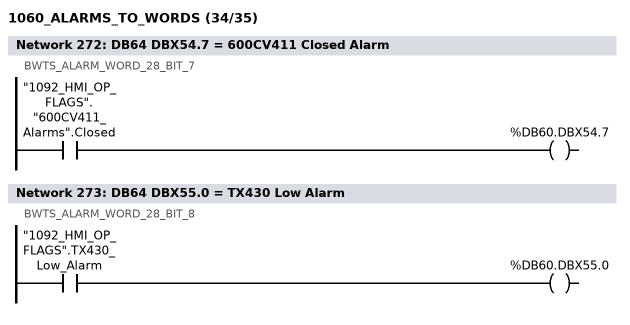
   RUNG wire#powerrail
      Contact( "1092_HMI_OP_FLAGS"."600CV411_Alarms".Closed )
      Coil( %DB60.DBX54.7 )
   END_RUNG
   // the same network as SCL:
   %DB60.DBX54.7 := "1092_HMI_OP_FLAGS"."600CV411_Alarms".Closed;
END_REGION

REGION Network 273: DB64 DBX55.0 = TX430 Low Alarm
   // BWTS_ALARM_WORD_28_BIT_8
   RUNG wire#powerrail
      Contact( "1092_HMI_OP_FLAGS".TX430_Low_Alarm )
      Coil( %DB60.DBX55.0 )
   END_RUNG
   // the same network as SCL:
   %DB60.DBX55.0 := "1092_HMI_OP_FLAGS".TX430_Low_Alarm;
END_REGION

REGION Network 275: Alarm Present
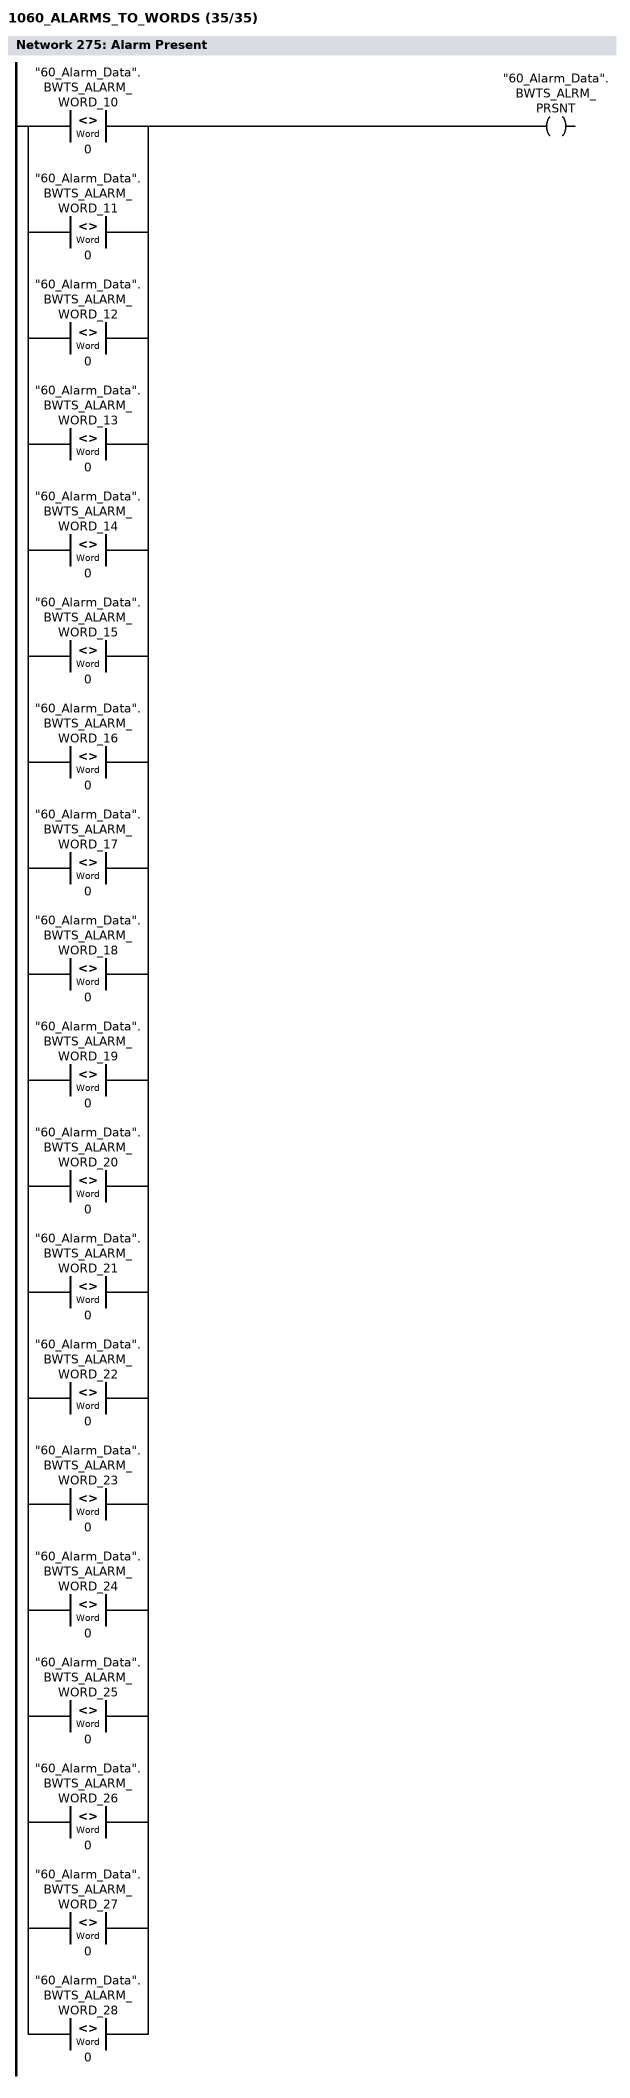
   RUNG wire#powerrail
      { S7_Templates := "SrcType := Word" } NE_Contact(in1 := "60_Alarm_Data".BWTS_ALARM_WORD_10, in2 := 0)
      wire#w1
      Coil( "60_Alarm_Data".BWTS_ALRM_PRSNT )
   END_RUNG
   RUNG wire#powerrail
      { S7_Templates := "SrcType := Word" } NE_Contact(in1 := "60_Alarm_Data".BWTS_ALARM_WORD_11, in2 := 0)
   END_RUNG wire#w1
   RUNG wire#powerrail
      { S7_Templates := "SrcType := Word" } NE_Contact(in1 := "60_Alarm_Data".BWTS_ALARM_WORD_12, in2 := 0)
   END_RUNG wire#w1
   RUNG wire#powerrail
      { S7_Templates := "SrcType := Word" } NE_Contact(in1 := "60_Alarm_Data".BWTS_ALARM_WORD_13, in2 := 0)
   END_RUNG wire#w1
   RUNG wire#powerrail
      { S7_Templates := "SrcType := Word" } NE_Contact(in1 := "60_Alarm_Data".BWTS_ALARM_WORD_14, in2 := 0)
   END_RUNG wire#w1
   RUNG wire#powerrail
      { S7_Templates := "SrcType := Word" } NE_Contact(in1 := "60_Alarm_Data".BWTS_ALARM_WORD_15, in2 := 0)
   END_RUNG wire#w1
   RUNG wire#powerrail
      { S7_Templates := "SrcType := Word" } NE_Contact(in1 := "60_Alarm_Data".BWTS_ALARM_WORD_16, in2 := 0)
   END_RUNG wire#w1
   RUNG wire#powerrail
      { S7_Templates := "SrcType := Word" } NE_Contact(in1 := "60_Alarm_Data".BWTS_ALARM_WORD_17, in2 := 0)
   END_RUNG wire#w1
   RUNG wire#powerrail
      { S7_Templates := "SrcType := Word" } NE_Contact(in1 := "60_Alarm_Data".BWTS_ALARM_WORD_18, in2 := 0)
   END_RUNG wire#w1
   RUNG wire#powerrail
      { S7_Templates := "SrcType := Word" } NE_Contact(in1 := "60_Alarm_Data".BWTS_ALARM_WORD_19, in2 := 0)
   END_RUNG wire#w1
   RUNG wire#powerrail
      { S7_Templates := "SrcType := Word" } NE_Contact(in1 := "60_Alarm_Data".BWTS_ALARM_WORD_20, in2 := 0)
   END_RUNG wire#w1
   RUNG wire#powerrail
      { S7_Templates := "SrcType := Word" } NE_Contact(in1 := "60_Alarm_Data".BWTS_ALARM_WORD_21, in2 := 0)
   END_RUNG wire#w1
   RUNG wire#powerrail
      { S7_Templates := "SrcType := Word" } NE_Contact(in1 := "60_Alarm_Data".BWTS_ALARM_WORD_22, in2 := 0)
   END_RUNG wire#w1
   RUNG wire#powerrail
      { S7_Templates := "SrcType := Word" } NE_Contact(in1 := "60_Alarm_Data".BWTS_ALARM_WORD_23, in2 := 0)
   END_RUNG wire#w1
   RUNG wire#powerrail
      { S7_Templates := "SrcType := Word" } NE_Contact(in1 := "60_Alarm_Data".BWTS_ALARM_WORD_24, in2 := 0)
   END_RUNG wire#w1
   RUNG wire#powerrail
      { S7_Templates := "SrcType := Word" } NE_Contact(in1 := "60_Alarm_Data".BWTS_ALARM_WORD_25, in2 := 0)
   END_RUNG wire#w1
   RUNG wire#powerrail
      { S7_Templates := "SrcType := Word" } NE_Contact(in1 := "60_Alarm_Data".BWTS_ALARM_WORD_26, in2 := 0)
   END_RUNG wire#w1
   RUNG wire#powerrail
      { S7_Templates := "SrcType := Word" } NE_Contact(in1 := "60_Alarm_Data".BWTS_ALARM_WORD_27, in2 := 0)
   END_RUNG wire#w1
   RUNG wire#powerrail
      { S7_Templates := "SrcType := Word" } NE_Contact(in1 := "60_Alarm_Data".BWTS_ALARM_WORD_28, in2 := 0)
   END_RUNG wire#w1
   // the same network as SCL:
   "60_Alarm_Data".BWTS_ALRM_PRSNT := ("60_Alarm_Data".BWTS_ALARM_WORD_10 <> 0) OR ("60_Alarm_Data".BWTS_ALARM_WORD_11 <> 0) OR ("60_Alarm_Data".BWTS_ALARM_WORD_12 <> 0) OR ("60_Alarm_Data".BWTS_ALARM_WORD_13 <> 0) OR ("60_Alarm_Data".BWTS_ALARM_WORD_14 <> 0) OR ("60_Alarm_Data".BWTS_ALARM_WORD_15 <> 0) OR ("60_Alarm_Data".BWTS_ALARM_WORD_16 <> 0) OR ("60_Alarm_Data".BWTS_ALARM_WORD_17 <> 0) OR ("60_Alarm_Data".BWTS_ALARM_WORD_18 <> 0) OR ("60_Alarm_Data".BWTS_ALARM_WORD_19 <> 0) OR ("60_Alarm_Data".BWTS_ALARM_WORD_20 <> 0) OR ("60_Alarm_Data".BWTS_ALARM_WORD_21 <> 0) OR ("60_Alarm_Data".BWTS_ALARM_WORD_22 <> 0) OR ("60_Alarm_Data".BWTS_ALARM_WORD_23 <> 0) OR ("60_Alarm_Data".BWTS_ALARM_WORD_24 <> 0) OR ("60_Alarm_Data".BWTS_ALARM_WORD_25 <> 0) OR ("60_Alarm_Data".BWTS_ALARM_WORD_26 <> 0) OR ("60_Alarm_Data".BWTS_ALARM_WORD_27 <> 0) OR ("60_Alarm_Data".BWTS_ALARM_WORD_28 <> 0);
END_REGION
END_FUNCTION

FUNCTION "1062_WARNINGS_TO_WORDS" : Void   // FC1062, LAD
TITLE = Warning Processing
{ S7_Optimized_Access := 'TRUE' }
AUTHOR : JRS
VERSION : 0.1
BEGIN

REGION Network 1: DB66 DBX18.0 = TX425/426 Tank 1 pH High Warning
   // BWTS_WARNING_WORD_10_BIT_0
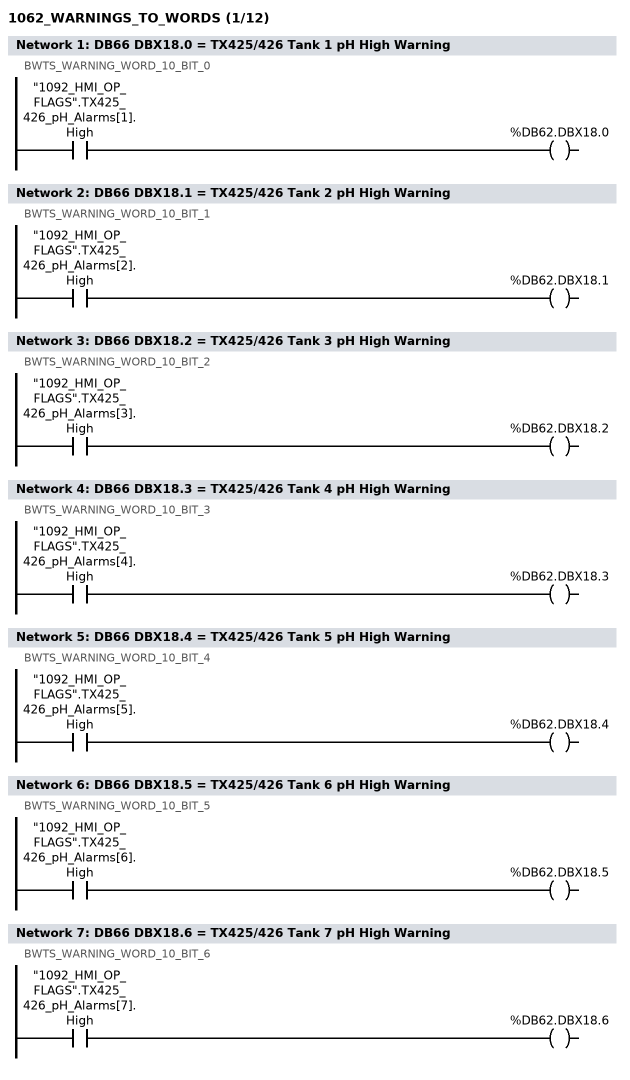
   RUNG wire#powerrail
      Contact( "1092_HMI_OP_FLAGS".TX425_426_pH_Alarms[1].High )
      Coil( %DB62.DBX18.0 )
   END_RUNG
   // the same network as SCL:
   %DB62.DBX18.0 := "1092_HMI_OP_FLAGS".TX425_426_pH_Alarms[1].High;
END_REGION

REGION Network 2: DB66 DBX18.1 = TX425/426 Tank 2 pH High Warning
   // BWTS_WARNING_WORD_10_BIT_1
   RUNG wire#powerrail
      Contact( "1092_HMI_OP_FLAGS".TX425_426_pH_Alarms[2].High )
      Coil( %DB62.DBX18.1 )
   END_RUNG
   // the same network as SCL:
   %DB62.DBX18.1 := "1092_HMI_OP_FLAGS".TX425_426_pH_Alarms[2].High;
END_REGION

REGION Network 3: DB66 DBX18.2 = TX425/426 Tank 3 pH High Warning
   // BWTS_WARNING_WORD_10_BIT_2
   RUNG wire#powerrail
      Contact( "1092_HMI_OP_FLAGS".TX425_426_pH_Alarms[3].High )
      Coil( %DB62.DBX18.2 )
   END_RUNG
   // the same network as SCL:
   %DB62.DBX18.2 := "1092_HMI_OP_FLAGS".TX425_426_pH_Alarms[3].High;
END_REGION

REGION Network 4: DB66 DBX18.3 = TX425/426 Tank 4 pH High Warning
   // BWTS_WARNING_WORD_10_BIT_3
   RUNG wire#powerrail
      Contact( "1092_HMI_OP_FLAGS".TX425_426_pH_Alarms[4].High )
      Coil( %DB62.DBX18.3 )
   END_RUNG
   // the same network as SCL:
   %DB62.DBX18.3 := "1092_HMI_OP_FLAGS".TX425_426_pH_Alarms[4].High;
END_REGION

REGION Network 5: DB66 DBX18.4 = TX425/426 Tank 5 pH High Warning
   // BWTS_WARNING_WORD_10_BIT_4
   RUNG wire#powerrail
      Contact( "1092_HMI_OP_FLAGS".TX425_426_pH_Alarms[5].High )
      Coil( %DB62.DBX18.4 )
   END_RUNG
   // the same network as SCL:
   %DB62.DBX18.4 := "1092_HMI_OP_FLAGS".TX425_426_pH_Alarms[5].High;
END_REGION

REGION Network 6: DB66 DBX18.5 = TX425/426 Tank 6 pH High Warning
   // BWTS_WARNING_WORD_10_BIT_5
   RUNG wire#powerrail
      Contact( "1092_HMI_OP_FLAGS".TX425_426_pH_Alarms[6].High )
      Coil( %DB62.DBX18.5 )
   END_RUNG
   // the same network as SCL:
   %DB62.DBX18.5 := "1092_HMI_OP_FLAGS".TX425_426_pH_Alarms[6].High;
END_REGION

REGION Network 7: DB66 DBX18.6 = TX425/426 Tank 7 pH High Warning
   // BWTS_WARNING_WORD_10_BIT_6
   RUNG wire#powerrail
      Contact( "1092_HMI_OP_FLAGS".TX425_426_pH_Alarms[7].High )
      Coil( %DB62.DBX18.6 )
   END_RUNG
   // the same network as SCL:
   %DB62.DBX18.6 := "1092_HMI_OP_FLAGS".TX425_426_pH_Alarms[7].High;
END_REGION

REGION Network 8: DB66 DBX18.7 = TX425/426 Tank 8 pH High Warning
   // BWTS_WARNING_WORD_10_BIT_7
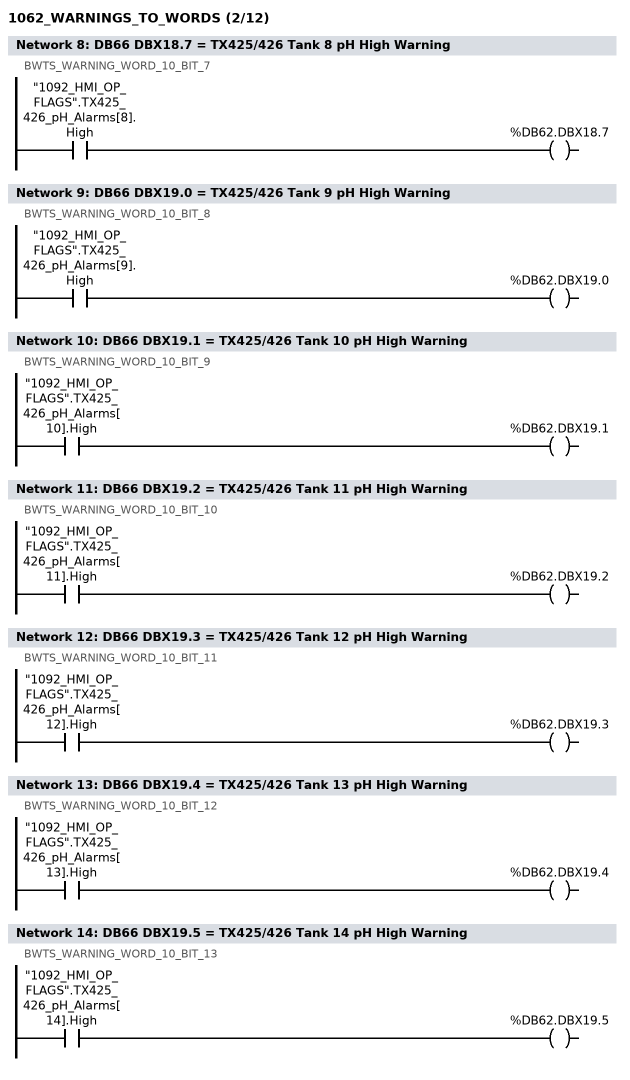
   RUNG wire#powerrail
      Contact( "1092_HMI_OP_FLAGS".TX425_426_pH_Alarms[8].High )
      Coil( %DB62.DBX18.7 )
   END_RUNG
   // the same network as SCL:
   %DB62.DBX18.7 := "1092_HMI_OP_FLAGS".TX425_426_pH_Alarms[8].High;
END_REGION

REGION Network 9: DB66 DBX19.0 = TX425/426 Tank 9 pH High Warning
   // BWTS_WARNING_WORD_10_BIT_8
   RUNG wire#powerrail
      Contact( "1092_HMI_OP_FLAGS".TX425_426_pH_Alarms[9].High )
      Coil( %DB62.DBX19.0 )
   END_RUNG
   // the same network as SCL:
   %DB62.DBX19.0 := "1092_HMI_OP_FLAGS".TX425_426_pH_Alarms[9].High;
END_REGION

REGION Network 10: DB66 DBX19.1 = TX425/426 Tank 10 pH High Warning
   // BWTS_WARNING_WORD_10_BIT_9
   RUNG wire#powerrail
      Contact( "1092_HMI_OP_FLAGS".TX425_426_pH_Alarms[10].High )
      Coil( %DB62.DBX19.1 )
   END_RUNG
   // the same network as SCL:
   %DB62.DBX19.1 := "1092_HMI_OP_FLAGS".TX425_426_pH_Alarms[10].High;
END_REGION

REGION Network 11: DB66 DBX19.2 = TX425/426 Tank 11 pH High Warning
   // BWTS_WARNING_WORD_10_BIT_10
   RUNG wire#powerrail
      Contact( "1092_HMI_OP_FLAGS".TX425_426_pH_Alarms[11].High )
      Coil( %DB62.DBX19.2 )
   END_RUNG
   // the same network as SCL:
   %DB62.DBX19.2 := "1092_HMI_OP_FLAGS".TX425_426_pH_Alarms[11].High;
END_REGION

REGION Network 12: DB66 DBX19.3 = TX425/426 Tank 12 pH High Warning
   // BWTS_WARNING_WORD_10_BIT_11
   RUNG wire#powerrail
      Contact( "1092_HMI_OP_FLAGS".TX425_426_pH_Alarms[12].High )
      Coil( %DB62.DBX19.3 )
   END_RUNG
   // the same network as SCL:
   %DB62.DBX19.3 := "1092_HMI_OP_FLAGS".TX425_426_pH_Alarms[12].High;
END_REGION

REGION Network 13: DB66 DBX19.4 = TX425/426 Tank 13 pH High Warning
   // BWTS_WARNING_WORD_10_BIT_12
   RUNG wire#powerrail
      Contact( "1092_HMI_OP_FLAGS".TX425_426_pH_Alarms[13].High )
      Coil( %DB62.DBX19.4 )
   END_RUNG
   // the same network as SCL:
   %DB62.DBX19.4 := "1092_HMI_OP_FLAGS".TX425_426_pH_Alarms[13].High;
END_REGION

REGION Network 14: DB66 DBX19.5 = TX425/426 Tank 14 pH High Warning
   // BWTS_WARNING_WORD_10_BIT_13
   RUNG wire#powerrail
      Contact( "1092_HMI_OP_FLAGS".TX425_426_pH_Alarms[14].High )
      Coil( %DB62.DBX19.5 )
   END_RUNG
   // the same network as SCL:
   %DB62.DBX19.5 := "1092_HMI_OP_FLAGS".TX425_426_pH_Alarms[14].High;
END_REGION

REGION Network 16: DB66 DBX20.0 = FIT417/418 Flow Tank 1 High Warning
   // BWTS_WARNING_WORD_11_BIT_0
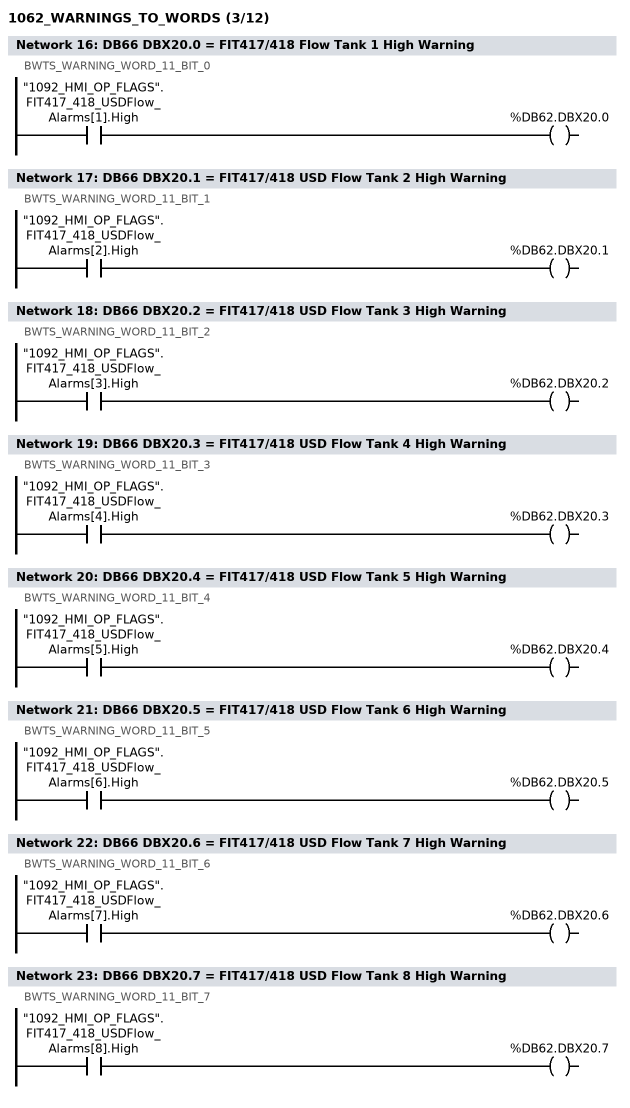
   RUNG wire#powerrail
      Contact( "1092_HMI_OP_FLAGS".FIT417_418_USDFlow_Alarms[1].High )
      Coil( %DB62.DBX20.0 )
   END_RUNG
   // the same network as SCL:
   %DB62.DBX20.0 := "1092_HMI_OP_FLAGS".FIT417_418_USDFlow_Alarms[1].High;
END_REGION

REGION Network 17: DB66 DBX20.1 = FIT417/418 USD Flow Tank 2 High Warning
   // BWTS_WARNING_WORD_11_BIT_1
   RUNG wire#powerrail
      Contact( "1092_HMI_OP_FLAGS".FIT417_418_USDFlow_Alarms[2].High )
      Coil( %DB62.DBX20.1 )
   END_RUNG
   // the same network as SCL:
   %DB62.DBX20.1 := "1092_HMI_OP_FLAGS".FIT417_418_USDFlow_Alarms[2].High;
END_REGION

REGION Network 18: DB66 DBX20.2 = FIT417/418 USD Flow Tank 3 High Warning
   // BWTS_WARNING_WORD_11_BIT_2
   RUNG wire#powerrail
      Contact( "1092_HMI_OP_FLAGS".FIT417_418_USDFlow_Alarms[3].High )
      Coil( %DB62.DBX20.2 )
   END_RUNG
   // the same network as SCL:
   %DB62.DBX20.2 := "1092_HMI_OP_FLAGS".FIT417_418_USDFlow_Alarms[3].High;
END_REGION

REGION Network 19: DB66 DBX20.3 = FIT417/418 USD Flow Tank 4 High Warning
   // BWTS_WARNING_WORD_11_BIT_3
   RUNG wire#powerrail
      Contact( "1092_HMI_OP_FLAGS".FIT417_418_USDFlow_Alarms[4].High )
      Coil( %DB62.DBX20.3 )
   END_RUNG
   // the same network as SCL:
   %DB62.DBX20.3 := "1092_HMI_OP_FLAGS".FIT417_418_USDFlow_Alarms[4].High;
END_REGION

REGION Network 20: DB66 DBX20.4 = FIT417/418 USD Flow Tank 5 High Warning
   // BWTS_WARNING_WORD_11_BIT_4
   RUNG wire#powerrail
      Contact( "1092_HMI_OP_FLAGS".FIT417_418_USDFlow_Alarms[5].High )
      Coil( %DB62.DBX20.4 )
   END_RUNG
   // the same network as SCL:
   %DB62.DBX20.4 := "1092_HMI_OP_FLAGS".FIT417_418_USDFlow_Alarms[5].High;
END_REGION

REGION Network 21: DB66 DBX20.5 = FIT417/418 USD Flow Tank 6 High Warning
   // BWTS_WARNING_WORD_11_BIT_5
   RUNG wire#powerrail
      Contact( "1092_HMI_OP_FLAGS".FIT417_418_USDFlow_Alarms[6].High )
      Coil( %DB62.DBX20.5 )
   END_RUNG
   // the same network as SCL:
   %DB62.DBX20.5 := "1092_HMI_OP_FLAGS".FIT417_418_USDFlow_Alarms[6].High;
END_REGION

REGION Network 22: DB66 DBX20.6 = FIT417/418 USD Flow Tank 7 High Warning
   // BWTS_WARNING_WORD_11_BIT_6
   RUNG wire#powerrail
      Contact( "1092_HMI_OP_FLAGS".FIT417_418_USDFlow_Alarms[7].High )
      Coil( %DB62.DBX20.6 )
   END_RUNG
   // the same network as SCL:
   %DB62.DBX20.6 := "1092_HMI_OP_FLAGS".FIT417_418_USDFlow_Alarms[7].High;
END_REGION

REGION Network 23: DB66 DBX20.7 = FIT417/418 USD Flow Tank 8 High Warning
   // BWTS_WARNING_WORD_11_BIT_7
   RUNG wire#powerrail
      Contact( "1092_HMI_OP_FLAGS".FIT417_418_USDFlow_Alarms[8].High )
      Coil( %DB62.DBX20.7 )
   END_RUNG
   // the same network as SCL:
   %DB62.DBX20.7 := "1092_HMI_OP_FLAGS".FIT417_418_USDFlow_Alarms[8].High;
END_REGION

REGION Network 24: DB66 DBX21.0 = FIT417/418 USD Flow Tank 9 High Warning
   // BWTS_WARNING_WORD_11_BIT_8
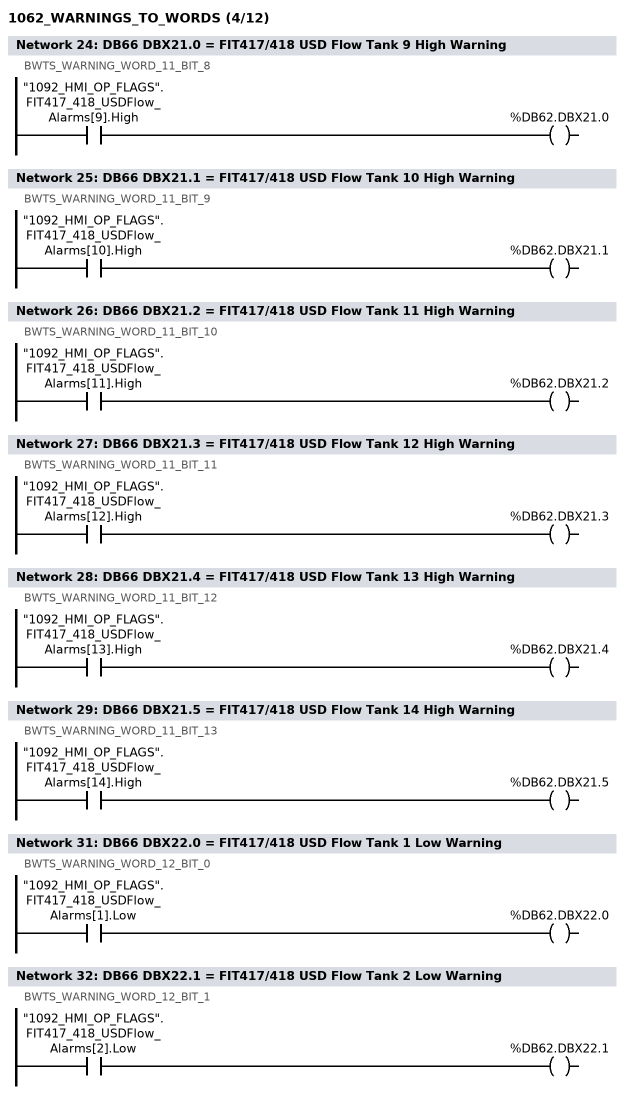
   RUNG wire#powerrail
      Contact( "1092_HMI_OP_FLAGS".FIT417_418_USDFlow_Alarms[9].High )
      Coil( %DB62.DBX21.0 )
   END_RUNG
   // the same network as SCL:
   %DB62.DBX21.0 := "1092_HMI_OP_FLAGS".FIT417_418_USDFlow_Alarms[9].High;
END_REGION

REGION Network 25: DB66 DBX21.1 = FIT417/418 USD Flow Tank 10 High Warning
   // BWTS_WARNING_WORD_11_BIT_9
   RUNG wire#powerrail
      Contact( "1092_HMI_OP_FLAGS".FIT417_418_USDFlow_Alarms[10].High )
      Coil( %DB62.DBX21.1 )
   END_RUNG
   // the same network as SCL:
   %DB62.DBX21.1 := "1092_HMI_OP_FLAGS".FIT417_418_USDFlow_Alarms[10].High;
END_REGION

REGION Network 26: DB66 DBX21.2 = FIT417/418 USD Flow Tank 11 High Warning
   // BWTS_WARNING_WORD_11_BIT_10
   RUNG wire#powerrail
      Contact( "1092_HMI_OP_FLAGS".FIT417_418_USDFlow_Alarms[11].High )
      Coil( %DB62.DBX21.2 )
   END_RUNG
   // the same network as SCL:
   %DB62.DBX21.2 := "1092_HMI_OP_FLAGS".FIT417_418_USDFlow_Alarms[11].High;
END_REGION

REGION Network 27: DB66 DBX21.3 = FIT417/418 USD Flow Tank 12 High Warning
   // BWTS_WARNING_WORD_11_BIT_11
   RUNG wire#powerrail
      Contact( "1092_HMI_OP_FLAGS".FIT417_418_USDFlow_Alarms[12].High )
      Coil( %DB62.DBX21.3 )
   END_RUNG
   // the same network as SCL:
   %DB62.DBX21.3 := "1092_HMI_OP_FLAGS".FIT417_418_USDFlow_Alarms[12].High;
END_REGION

REGION Network 28: DB66 DBX21.4 = FIT417/418 USD Flow Tank 13 High Warning
   // BWTS_WARNING_WORD_11_BIT_12
   RUNG wire#powerrail
      Contact( "1092_HMI_OP_FLAGS".FIT417_418_USDFlow_Alarms[13].High )
      Coil( %DB62.DBX21.4 )
   END_RUNG
   // the same network as SCL:
   %DB62.DBX21.4 := "1092_HMI_OP_FLAGS".FIT417_418_USDFlow_Alarms[13].High;
END_REGION

REGION Network 29: DB66 DBX21.5 = FIT417/418 USD Flow Tank 14 High Warning
   // BWTS_WARNING_WORD_11_BIT_13
   RUNG wire#powerrail
      Contact( "1092_HMI_OP_FLAGS".FIT417_418_USDFlow_Alarms[14].High )
      Coil( %DB62.DBX21.5 )
   END_RUNG
   // the same network as SCL:
   %DB62.DBX21.5 := "1092_HMI_OP_FLAGS".FIT417_418_USDFlow_Alarms[14].High;
END_REGION

REGION Network 31: DB66 DBX22.0 = FIT417/418 USD Flow Tank 1 Low Warning
   // BWTS_WARNING_WORD_12_BIT_0
   RUNG wire#powerrail
      Contact( "1092_HMI_OP_FLAGS".FIT417_418_USDFlow_Alarms[1].Low )
      Coil( %DB62.DBX22.0 )
   END_RUNG
   // the same network as SCL:
   %DB62.DBX22.0 := "1092_HMI_OP_FLAGS".FIT417_418_USDFlow_Alarms[1].Low;
END_REGION

REGION Network 32: DB66 DBX22.1 = FIT417/418 USD Flow Tank 2 Low Warning
   // BWTS_WARNING_WORD_12_BIT_1
   RUNG wire#powerrail
      Contact( "1092_HMI_OP_FLAGS".FIT417_418_USDFlow_Alarms[2].Low )
      Coil( %DB62.DBX22.1 )
   END_RUNG
   // the same network as SCL:
   %DB62.DBX22.1 := "1092_HMI_OP_FLAGS".FIT417_418_USDFlow_Alarms[2].Low;
END_REGION

REGION Network 33: DB66 DBX22.2 = FIT417/418 USD Flow Tank 3 Low Warning
   // BWTS_WARNING_WORD_12_BIT_2
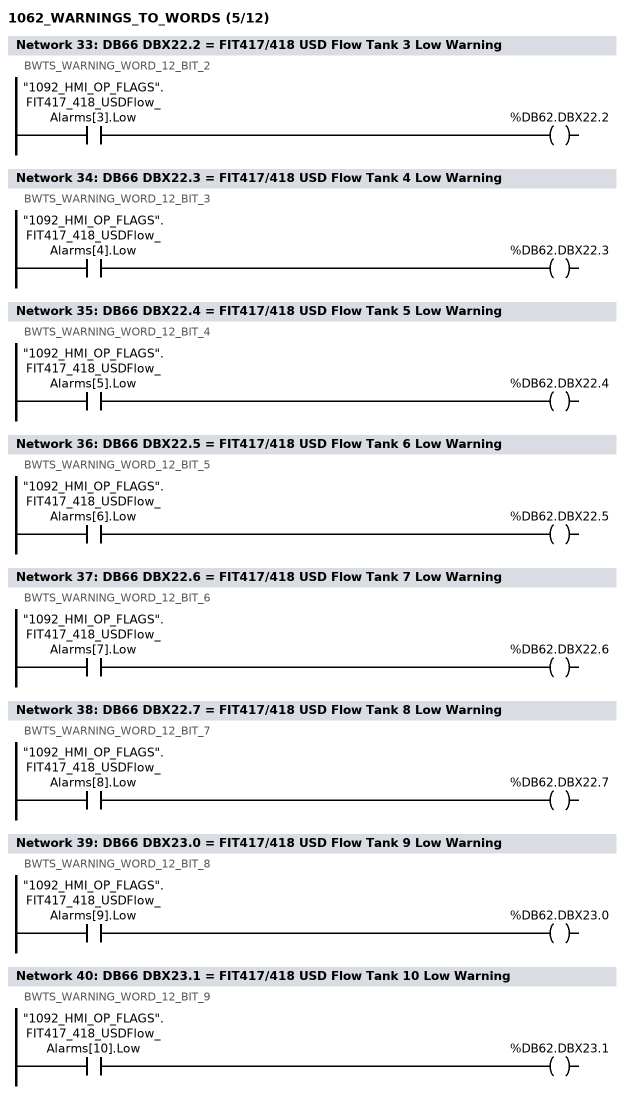
   RUNG wire#powerrail
      Contact( "1092_HMI_OP_FLAGS".FIT417_418_USDFlow_Alarms[3].Low )
      Coil( %DB62.DBX22.2 )
   END_RUNG
   // the same network as SCL:
   %DB62.DBX22.2 := "1092_HMI_OP_FLAGS".FIT417_418_USDFlow_Alarms[3].Low;
END_REGION

REGION Network 34: DB66 DBX22.3 = FIT417/418 USD Flow Tank 4 Low Warning
   // BWTS_WARNING_WORD_12_BIT_3
   RUNG wire#powerrail
      Contact( "1092_HMI_OP_FLAGS".FIT417_418_USDFlow_Alarms[4].Low )
      Coil( %DB62.DBX22.3 )
   END_RUNG
   // the same network as SCL:
   %DB62.DBX22.3 := "1092_HMI_OP_FLAGS".FIT417_418_USDFlow_Alarms[4].Low;
END_REGION

REGION Network 35: DB66 DBX22.4 = FIT417/418 USD Flow Tank 5 Low Warning
   // BWTS_WARNING_WORD_12_BIT_4
   RUNG wire#powerrail
      Contact( "1092_HMI_OP_FLAGS".FIT417_418_USDFlow_Alarms[5].Low )
      Coil( %DB62.DBX22.4 )
   END_RUNG
   // the same network as SCL:
   %DB62.DBX22.4 := "1092_HMI_OP_FLAGS".FIT417_418_USDFlow_Alarms[5].Low;
END_REGION

REGION Network 36: DB66 DBX22.5 = FIT417/418 USD Flow Tank 6 Low Warning
   // BWTS_WARNING_WORD_12_BIT_5
   RUNG wire#powerrail
      Contact( "1092_HMI_OP_FLAGS".FIT417_418_USDFlow_Alarms[6].Low )
      Coil( %DB62.DBX22.5 )
   END_RUNG
   // the same network as SCL:
   %DB62.DBX22.5 := "1092_HMI_OP_FLAGS".FIT417_418_USDFlow_Alarms[6].Low;
END_REGION

REGION Network 37: DB66 DBX22.6 = FIT417/418 USD Flow Tank 7 Low Warning
   // BWTS_WARNING_WORD_12_BIT_6
   RUNG wire#powerrail
      Contact( "1092_HMI_OP_FLAGS".FIT417_418_USDFlow_Alarms[7].Low )
      Coil( %DB62.DBX22.6 )
   END_RUNG
   // the same network as SCL:
   %DB62.DBX22.6 := "1092_HMI_OP_FLAGS".FIT417_418_USDFlow_Alarms[7].Low;
END_REGION

REGION Network 38: DB66 DBX22.7 = FIT417/418 USD Flow Tank 8 Low Warning
   // BWTS_WARNING_WORD_12_BIT_7
   RUNG wire#powerrail
      Contact( "1092_HMI_OP_FLAGS".FIT417_418_USDFlow_Alarms[8].Low )
      Coil( %DB62.DBX22.7 )
   END_RUNG
   // the same network as SCL:
   %DB62.DBX22.7 := "1092_HMI_OP_FLAGS".FIT417_418_USDFlow_Alarms[8].Low;
END_REGION

REGION Network 39: DB66 DBX23.0 = FIT417/418 USD Flow Tank 9 Low Warning
   // BWTS_WARNING_WORD_12_BIT_8
   RUNG wire#powerrail
      Contact( "1092_HMI_OP_FLAGS".FIT417_418_USDFlow_Alarms[9].Low )
      Coil( %DB62.DBX23.0 )
   END_RUNG
   // the same network as SCL:
   %DB62.DBX23.0 := "1092_HMI_OP_FLAGS".FIT417_418_USDFlow_Alarms[9].Low;
END_REGION

REGION Network 40: DB66 DBX23.1 = FIT417/418 USD Flow Tank 10 Low Warning
   // BWTS_WARNING_WORD_12_BIT_9
   RUNG wire#powerrail
      Contact( "1092_HMI_OP_FLAGS".FIT417_418_USDFlow_Alarms[10].Low )
      Coil( %DB62.DBX23.1 )
   END_RUNG
   // the same network as SCL:
   %DB62.DBX23.1 := "1092_HMI_OP_FLAGS".FIT417_418_USDFlow_Alarms[10].Low;
END_REGION

REGION Network 41: DB66 DBX23.2 = FIT417/418 USD Flow Tank 11 Low Warning
   // BWTS_WARNING_WORD_12_BIT_10
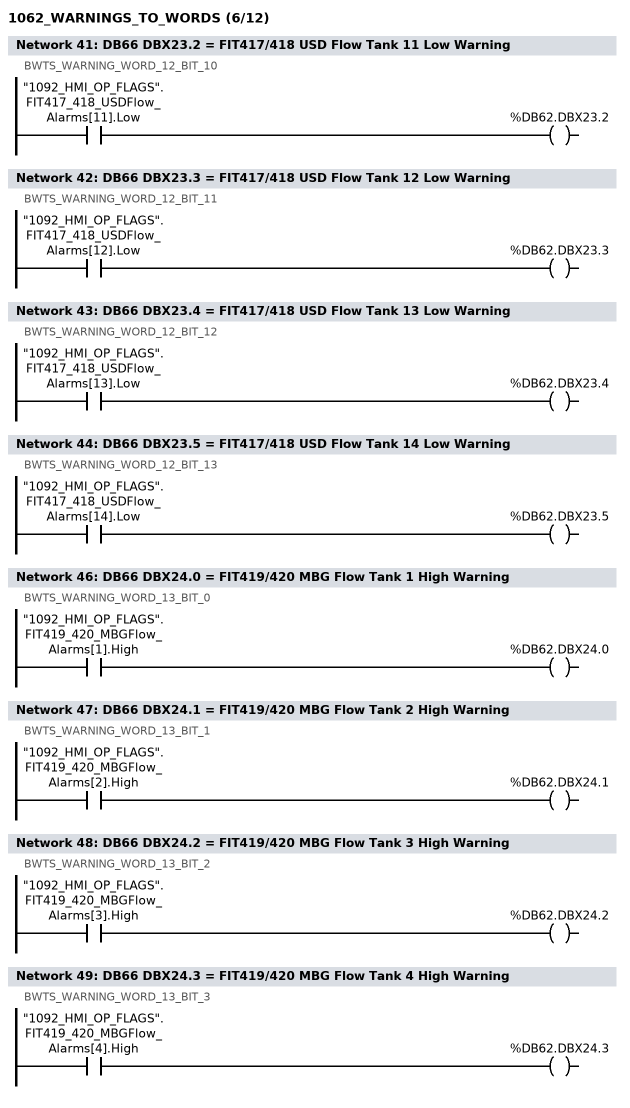
   RUNG wire#powerrail
      Contact( "1092_HMI_OP_FLAGS".FIT417_418_USDFlow_Alarms[11].Low )
      Coil( %DB62.DBX23.2 )
   END_RUNG
   // the same network as SCL:
   %DB62.DBX23.2 := "1092_HMI_OP_FLAGS".FIT417_418_USDFlow_Alarms[11].Low;
END_REGION

REGION Network 42: DB66 DBX23.3 = FIT417/418 USD Flow Tank 12 Low Warning
   // BWTS_WARNING_WORD_12_BIT_11
   RUNG wire#powerrail
      Contact( "1092_HMI_OP_FLAGS".FIT417_418_USDFlow_Alarms[12].Low )
      Coil( %DB62.DBX23.3 )
   END_RUNG
   // the same network as SCL:
   %DB62.DBX23.3 := "1092_HMI_OP_FLAGS".FIT417_418_USDFlow_Alarms[12].Low;
END_REGION

REGION Network 43: DB66 DBX23.4 = FIT417/418 USD Flow Tank 13 Low Warning
   // BWTS_WARNING_WORD_12_BIT_12
   RUNG wire#powerrail
      Contact( "1092_HMI_OP_FLAGS".FIT417_418_USDFlow_Alarms[13].Low )
      Coil( %DB62.DBX23.4 )
   END_RUNG
   // the same network as SCL:
   %DB62.DBX23.4 := "1092_HMI_OP_FLAGS".FIT417_418_USDFlow_Alarms[13].Low;
END_REGION

REGION Network 44: DB66 DBX23.5 = FIT417/418 USD Flow Tank 14 Low Warning
   // BWTS_WARNING_WORD_12_BIT_13
   RUNG wire#powerrail
      Contact( "1092_HMI_OP_FLAGS".FIT417_418_USDFlow_Alarms[14].Low )
      Coil( %DB62.DBX23.5 )
   END_RUNG
   // the same network as SCL:
   %DB62.DBX23.5 := "1092_HMI_OP_FLAGS".FIT417_418_USDFlow_Alarms[14].Low;
END_REGION

REGION Network 46: DB66 DBX24.0 = FIT419/420 MBG Flow Tank 1 High Warning
   // BWTS_WARNING_WORD_13_BIT_0
   RUNG wire#powerrail
      Contact( "1092_HMI_OP_FLAGS".FIT419_420_MBGFlow_Alarms[1].High )
      Coil( %DB62.DBX24.0 )
   END_RUNG
   // the same network as SCL:
   %DB62.DBX24.0 := "1092_HMI_OP_FLAGS".FIT419_420_MBGFlow_Alarms[1].High;
END_REGION

REGION Network 47: DB66 DBX24.1 = FIT419/420 MBG Flow Tank 2 High Warning
   // BWTS_WARNING_WORD_13_BIT_1
   RUNG wire#powerrail
      Contact( "1092_HMI_OP_FLAGS".FIT419_420_MBGFlow_Alarms[2].High )
      Coil( %DB62.DBX24.1 )
   END_RUNG
   // the same network as SCL:
   %DB62.DBX24.1 := "1092_HMI_OP_FLAGS".FIT419_420_MBGFlow_Alarms[2].High;
END_REGION

REGION Network 48: DB66 DBX24.2 = FIT419/420 MBG Flow Tank 3 High Warning
   // BWTS_WARNING_WORD_13_BIT_2
   RUNG wire#powerrail
      Contact( "1092_HMI_OP_FLAGS".FIT419_420_MBGFlow_Alarms[3].High )
      Coil( %DB62.DBX24.2 )
   END_RUNG
   // the same network as SCL:
   %DB62.DBX24.2 := "1092_HMI_OP_FLAGS".FIT419_420_MBGFlow_Alarms[3].High;
END_REGION

REGION Network 49: DB66 DBX24.3 = FIT419/420 MBG Flow Tank 4 High Warning
   // BWTS_WARNING_WORD_13_BIT_3
   RUNG wire#powerrail
      Contact( "1092_HMI_OP_FLAGS".FIT419_420_MBGFlow_Alarms[4].High )
      Coil( %DB62.DBX24.3 )
   END_RUNG
   // the same network as SCL:
   %DB62.DBX24.3 := "1092_HMI_OP_FLAGS".FIT419_420_MBGFlow_Alarms[4].High;
END_REGION

REGION Network 50: DB66 DBX24.4 = FIT419/420 MBG Flow Tank 5 High Warning
   // BWTS_WARNING_WORD_13_BIT_4
